   694: 'Spare_Fault_694', class No Acknowledgement, trigger "DB302_HMI_Faults_Carrier10_Faults_3" bit 5
   695: 'Spare_Fault_695', class No Acknowledgement, trigger "DB302_HMI_Faults_Carrier10_Faults_3" bit 6
   696: 'Spare_Fault_696', class No Acknowledgement, trigger "DB302_HMI_Faults_Carrier10_Faults_3" bit 7
   697: 'Spare_Fault_697', class No Acknowledgement, trigger "DB302_HMI_Faults_Carrier10_Faults_3" bit 8
   698: 'Spare_Fault_698', class No Acknowledgement, trigger "DB302_HMI_Faults_Carrier10_Faults_3" bit 9
   699: 'Spare_Fault_699', class No Acknowledgement, trigger "DB302_HMI_Faults_Carrier10_Faults_3" bit 10
   700: 'Spare_Fault_700', class No Acknowledgement, trigger "DB302_HMI_Faults_Carrier10_Faults_3" bit 11
   701: 'Spare_Fault_701', class No Acknowledgement, trigger "DB302_HMI_Faults_Carrier10_Faults_3" bit 12
   702: 'Spare_Fault_702', class No Acknowledgement, trigger "DB302_HMI_Faults_Carrier10_Faults_3" bit 13
   703: 'Spare_Fault_703', class No Acknowledgement, trigger "DB302_HMI_Faults_Carrier10_Faults_3" bit 14
   704: 'Spare_Fault_704', class No Acknowledgement, trigger "DB302_HMI_Faults_Carrier10_Faults_3" bit 15
   705: 'Carrier 11 Disconnect Open Power Fault DI11.0', class No Acknowledgement, trigger "DB302_HMI_Faults_Carrier11_Faults_0" bit 0
   706: 'Carrier 11 Drive Profinet Comm Fault', class No Acknowledgement, trigger "DB302_HMI_Faults_Carrier11_Faults_0" bit 1
   707: 'Carrier 11 Production Stop Not Reset', class No Acknowledgement, trigger "DB302_HMI_Faults_Carrier11_Faults_0" bit 2
   708: 'Carrier 11 CB02122 Tripped', class No Acknowledgement, trigger "DB302_HMI_Faults_Carrier11_Faults_0" bit 3
   709: 'Carrier 11 CB02123 Tripped', class No Acknowledgement, trigger "DB302_HMI_Faults_Carrier11_Faults_0" bit 4
   710: 'Carrier 11 AUX1 CB Tripped', class No Acknowledgement, trigger "DB302_HMI_Faults_Carrier11_Faults_0" bit 5
   711: 'Carrier 11 AUX2 CB Tripped', class No Acknowledgement, trigger "DB302_HMI_Faults_Carrier11_Faults_0" bit 6
   712: 'Carrier 11 PLC Not Communicating', class No Acknowledgement, trigger "DB302_HMI_Faults_Carrier11_Faults_0" bit 7
   713: 'Carrier 11 Safe Input Card Fault', class No Acknowledgement, trigger "DB302_HMI_Faults_Carrier11_Faults_0" bit 8
   714: 'Carrier 11 Safe Output Card Fault', class No Acknowledgement, trigger "DB302_HMI_Faults_Carrier11_Faults_0" bit 9
   715: 'Carrier 11 Standard Input Card Fault', class No Acknowledgement, trigger "DB302_HMI_Faults_Carrier11_Faults_0" bit 10
   716: 'Carrier 11 Standard Output Card Fault', class No Acknowledgement, trigger "DB302_HMI_Faults_Carrier11_Faults_0" bit 11
   717: 'Carrier 11 Encoder Position Fault', class No Acknowledgement, trigger "DB302_HMI_Faults_Carrier11_Faults_0" bit 12
   718: 'Carrier 11 Encoder Internal Error', class No Acknowledgement, trigger "DB302_HMI_Faults_Carrier11_Faults_0" bit 13
   719: 'Carrier 11 Encoder Comm Fault', class No Acknowledgement, trigger "DB302_HMI_Faults_Carrier11_Faults_0" bit 14
   720: 'Carrier 11 HMI Comm Fault', class No Acknowledgement, trigger "DB302_HMI_Faults_Carrier11_Faults_0" bit 15
   721: 'Carrier 11 Crash Detection Fault', class No Acknowledgement, trigger "DB302_HMI_Faults_Carrier11_Faults_1" bit 0
   722: 'Carrier 11 Carrier Number Invalid', class No Acknowledgement, trigger "DB302_HMI_Faults_Carrier11_Faults_1" bit 1
   723: 'Carrier 11 Drive: PROFINET configuration error', class No Acknowledgement, trigger "DB302_HMI_Faults_Carrier11_Faults_1" bit 2
   724: 'Carrier 11 Drive: Error internal communications', class No Acknowledgement, trigger "DB302_HMI_Faults_Carrier11_Faults_1" bit 3
   725: 'Carrier 11 Drive: Motor overtemperature', class No Acknowledgement, trigger "DB302_HMI_Faults_Carrier11_Faults_1" bit 4
   726: 'Carrier 11 Drive: Motor overcurrent', class No Acknowledgement, trigger "DB302_HMI_Faults_Carrier11_Faults_1" bit 5
   727: 'Carrier 11 Drive: Infeed or power unit not ready', class No Acknowledgement, trigger "DB302_HMI_Faults_Carrier11_Faults_1" bit 6
   728: 'Carrier 11 Drive: Short-circuit/ground fault detected', class No Acknowledgement, trigger "DB302_HMI_Faults_Carrier11_Faults_1" bit 7
   729: 'Carrier 11 Drive: PROFINET Setpoint timeout', class No Acknowledgement, trigger "DB302_HMI_Faults_Carrier11_Faults_1" bit 8
   730: 'Carrier 11 Power unit: Overcurrent', class No Acknowledgement, trigger "DB302_HMI_Faults_Carrier11_Faults_1" bit 9
   731: 'Carrier 11 Power unit: DC link voltage overvoltage', class No Acknowledgement, trigger "DB302_HMI_Faults_Carrier11_Faults_1" bit 10
   732: 'Carrier 11 Power unit: DC link voltage undervoltage', class No Acknowledgement, trigger "DB302_HMI_Faults_Carrier11_Faults_1" bit 11
   733: 'Carrier 11 Power unit: Line phase failure in main circuit', class No Acknowledgement, trigger "DB302_HMI_Faults_Carrier11_Faults_1" bit 12
   734: 'Carrier 11 Power unit: Phase failure motor cable', class No Acknowledgement, trigger "DB302_HMI_Faults_Carrier11_Faults_1" bit 13
   735: 'Carrier 11 Power unit: Ground fault', class No Acknowledgement, trigger "DB302_HMI_Faults_Carrier11_Faults_1" bit 14
   736: 'Spare_Fault_736', class No Acknowledgement, trigger "DB302_HMI_Faults_Carrier11_Faults_1" bit 15
   737: 'Carrier 11 Motion Off Fault', class No Acknowledgement, trigger "DB302_HMI_Faults_Carrier11_Faults_2" bit 0
   738: 'Carrier 11 Motion On Fault', class No Acknowledgement, trigger "DB302_HMI_Faults_Carrier11_Faults_2" bit 1
   739: 'Carrier 11 Spacing Fault', class No Acknowledgement, trigger "DB302_HMI_Faults_Carrier11_Faults_2" bit 2
   740: 'Carrier 11 Duplicate Carrier Number Fault', class No Acknowledgement, trigger "DB302_HMI_Faults_Carrier11_Faults_2" bit 3
   741: 'Spare_Fault_741', class No Acknowledgement, trigger "DB302_HMI_Faults_Carrier11_Faults_2" bit 4
   742: 'Spare_Fault_742', class No Acknowledgement, trigger "DB302_HMI_Faults_Carrier11_Faults_2" bit 5
   743: 'Spare_Fault_743', class No Acknowledgement, trigger "DB302_HMI_Faults_Carrier11_Faults_2" bit 6
   744: 'Spare_Fault_744', class No Acknowledgement, trigger "DB302_HMI_Faults_Carrier11_Faults_2" bit 7
   745: 'Spare_Fault_745', class No Acknowledgement, trigger "DB302_HMI_Faults_Carrier11_Faults_2" bit 8
   746: 'Spare_Fault_746', class No Acknowledgement, trigger "DB302_HMI_Faults_Carrier11_Faults_2" bit 9
   747: 'Spare_Fault_747', class No Acknowledgement, trigger "DB302_HMI_Faults_Carrier11_Faults_2" bit 10
   748: 'Spare_Fault_748', class No Acknowledgement, trigger "DB302_HMI_Faults_Carrier11_Faults_2" bit 11
   749: 'Spare_Fault_749', class No Acknowledgement, trigger "DB302_HMI_Faults_Carrier11_Faults_2" bit 12
   750: 'Spare_Fault_750', class No Acknowledgement, trigger "DB302_HMI_Faults_Carrier11_Faults_2" bit 13
   751: 'Spare_Fault_751', class No Acknowledgement, trigger "DB302_HMI_Faults_Carrier11_Faults_2" bit 14
   752: 'Spare_Fault_752', class No Acknowledgement, trigger "DB302_HMI_Faults_Carrier11_Faults_2" bit 15
   753: 'Spare_Fault_753', class No Acknowledgement, trigger "DB302_HMI_Faults_Carrier11_Faults_3" bit 0
   754: 'Spare_Fault_754', class No Acknowledgement, trigger "DB302_HMI_Faults_Carrier11_Faults_3" bit 1
   755: 'Spare_Fault_755', class No Acknowledgement, trigger "DB302_HMI_Faults_Carrier11_Faults_3" bit 2
   756: 'Spare_Fault_756', class No Acknowledgement, trigger "DB302_HMI_Faults_Carrier11_Faults_3" bit 3
   757: 'Spare_Fault_757', class No Acknowledgement, trigger "DB302_HMI_Faults_Carrier11_Faults_3" bit 4
   758: 'Spare_Fault_758', class No Acknowledgement, trigger "DB302_HMI_Faults_Carrier11_Faults_3" bit 5
   759: 'Spare_Fault_759', class No Acknowledgement, trigger "DB302_HMI_Faults_Carrier11_Faults_3" bit 6
   760: 'Spare_Fault_760', class No Acknowledgement, trigger "DB302_HMI_Faults_Carrier11_Faults_3" bit 7
   761: 'Spare_Fault_761', class No Acknowledgement, trigger "DB302_HMI_Faults_Carrier11_Faults_3" bit 8
   762: 'Spare_Fault_762', class No Acknowledgement, trigger "DB302_HMI_Faults_Carrier11_Faults_3" bit 9
   763: 'Spare_Fault_763', class No Acknowledgement, trigger "DB302_HMI_Faults_Carrier11_Faults_3" bit 10
   764: 'Spare_Fault_764', class No Acknowledgement, trigger "DB302_HMI_Faults_Carrier11_Faults_3" bit 11
   765: 'Spare_Fault_765', class No Acknowledgement, trigger "DB302_HMI_Faults_Carrier11_Faults_3" bit 12
   766: 'Spare_Fault_766', class No Acknowledgement, trigger "DB302_HMI_Faults_Carrier11_Faults_3" bit 13
   767: 'Spare_Fault_767', class No Acknowledgement, trigger "DB302_HMI_Faults_Carrier11_Faults_3" bit 14
   768: 'Spare_Fault_768', class No Acknowledgement, trigger "DB302_HMI_Faults_Carrier11_Faults_3" bit 15
   769: 'Carrier 12 Disconnect Open Power Fault DI11.0', class No Acknowledgement, trigger "DB302_HMI_Faults_Carrier12_Faults_0" bit 0
   770: 'Carrier 12 Drive Profinet Comm Fault', class No Acknowledgement, trigger "DB302_HMI_Faults_Carrier12_Faults_0" bit 1
   771: 'Carrier 12 Production Stop Not Reset', class No Acknowledgement, trigger "DB302_HMI_Faults_Carrier12_Faults_0" bit 2
   772: 'Carrier 12 CB02122 Tripped', class No Acknowledgement, trigger "DB302_HMI_Faults_Carrier12_Faults_0" bit 3
   773: 'Carrier 12 CB02123 Tripped', class No Acknowledgement, trigger "DB302_HMI_Faults_Carrier12_Faults_0" bit 4
   774: 'Carrier 12 AUX1 CB Tripped', class No Acknowledgement, trigger "DB302_HMI_Faults_Carrier12_Faults_0" bit 5
   775: 'Carrier 12 AUX2 CB Tripped', class No Acknowledgement, trigger "DB302_HMI_Faults_Carrier12_Faults_0" bit 6
   776: 'Carrier 12 PLC Not Communicating', class No Acknowledgement, trigger "DB302_HMI_Faults_Carrier12_Faults_0" bit 7
   777: 'Carrier 12 Safe Input Card Fault', class No Acknowledgement, trigger "DB302_HMI_Faults_Carrier12_Faults_0" bit 8
   778: 'Carrier 12 Safe Output Card Fault', class No Acknowledgement, trigger "DB302_HMI_Faults_Carrier12_Faults_0" bit 9
   779: 'Carrier 12 Standard Input Card Fault', class No Acknowledgement, trigger "DB302_HMI_Faults_Carrier12_Faults_0" bit 10
   780: 'Carrier 12 Standard Output Card Fault', class No Acknowledgement, trigger "DB302_HMI_Faults_Carrier12_Faults_0" bit 11
   781: 'Carrier 12 Encoder Position Fault', class No Acknowledgement, trigger "DB302_HMI_Faults_Carrier12_Faults_0" bit 12
   782: 'Carrier 12 Encoder Internal Error', class No Acknowledgement, trigger "DB302_HMI_Faults_Carrier12_Faults_0" bit 13
   783: 'Carrier 12 Encoder Comm Fault', class No Acknowledgement, trigger "DB302_HMI_Faults_Carrier12_Faults_0" bit 14
   784: 'Carrier 12 HMI Comm Fault', class No Acknowledgement, trigger "DB302_HMI_Faults_Carrier12_Faults_0" bit 15
   785: 'Carrier 12 Crash Detection Fault', class No Acknowledgement, trigger "DB302_HMI_Faults_Carrier12_Faults_1" bit 0
   786: 'Carrier 12 Carrier Number Invalid', class No Acknowledgement, trigger "DB302_HMI_Faults_Carrier12_Faults_1" bit 1
   787: 'Carrier 12 Drive: PROFINET configuration error', class No Acknowledgement, trigger "DB302_HMI_Faults_Carrier12_Faults_1" bit 2
   788: 'Carrier 12 Drive: Error internal communications', class No Acknowledgement, trigger "DB302_HMI_Faults_Carrier12_Faults_1" bit 3
   789: 'Carrier 12 Drive: Motor overtemperature', class No Acknowledgement, trigger "DB302_HMI_Faults_Carrier12_Faults_1" bit 4
   790: 'Carrier 12 Drive: Motor overcurrent', class No Acknowledgement, trigger "DB302_HMI_Faults_Carrier12_Faults_1" bit 5
   791: 'Carrier 12 Drive: Infeed or power unit not ready', class No Acknowledgement, trigger "DB302_HMI_Faults_Carrier12_Faults_1" bit 6
   792: 'Carrier 12 Drive: Short-circuit/ground fault detected', class No Acknowledgement, trigger "DB302_HMI_Faults_Carrier12_Faults_1" bit 7
   793: 'Carrier 12 Drive: PROFINET Setpoint timeout', class No Acknowledgement, trigger "DB302_HMI_Faults_Carrier12_Faults_1" bit 8
   794: 'Carrier 12 Power unit: Overcurrent', class No Acknowledgement, trigger "DB302_HMI_Faults_Carrier12_Faults_1" bit 9
   795: 'Carrier 12 Power unit: DC link voltage overvoltage', class No Acknowledgement, trigger "DB302_HMI_Faults_Carrier12_Faults_1" bit 10
   796: 'Carrier 12 Power unit: DC link voltage undervoltage', class No Acknowledgement, trigger "DB302_HMI_Faults_Carrier12_Faults_1" bit 11
   797: 'Carrier 12 Power unit: Line phase failure in main circuit', class No Acknowledgement, trigger "DB302_HMI_Faults_Carrier12_Faults_1" bit 12
   798: 'Carrier 12 Power unit: Phase failure motor cable', class No Acknowledgement, trigger "DB302_HMI_Faults_Carrier12_Faults_1" bit 13
   799: 'Carrier 12 Power unit: Ground fault', class No Acknowledgement, trigger "DB302_HMI_Faults_Carrier12_Faults_1" bit 14
   800: 'Spare_Fault_800', class No Acknowledgement, trigger "DB302_HMI_Faults_Carrier12_Faults_1" bit 15
   801: 'Carrier 12 Motion Off Fault', class No Acknowledgement, trigger "DB302_HMI_Faults_Carrier12_Faults_2" bit 0
   802: 'Carrier 12 Motion On Fault', class No Acknowledgement, trigger "DB302_HMI_Faults_Carrier12_Faults_2" bit 1
   803: 'Carrier 12 Spacing Fault', class No Acknowledgement, trigger "DB302_HMI_Faults_Carrier12_Faults_2" bit 2
   804: 'Carrier 12 Duplicate Carrier Number Fault', class No Acknowledgement, trigger "DB302_HMI_Faults_Carrier12_Faults_2" bit 3
   805: 'Spare_Fault_805', class No Acknowledgement, trigger "DB302_HMI_Faults_Carrier12_Faults_2" bit 4
   806: 'Spare_Fault_806', class No Acknowledgement, trigger "DB302_HMI_Faults_Carrier12_Faults_2" bit 5
   807: 'Spare_Fault_807', class No Acknowledgement, trigger "DB302_HMI_Faults_Carrier12_Faults_2" bit 6
   808: 'Spare_Fault_808', class No Acknowledgement, trigger "DB302_HMI_Faults_Carrier12_Faults_2" bit 7
   809: 'Spare_Fault_809', class No Acknowledgement, trigger "DB302_HMI_Faults_Carrier12_Faults_2" bit 8
   810: 'Spare_Fault_810', class No Acknowledgement, trigger "DB302_HMI_Faults_Carrier12_Faults_2" bit 9
   811: 'Spare_Fault_811', class No Acknowledgement, trigger "DB302_HMI_Faults_Carrier12_Faults_2" bit 10
   812: 'Spare_Fault_812', class No Acknowledgement, trigger "DB302_HMI_Faults_Carrier12_Faults_2" bit 11
   813: 'Spare_Fault_813', class No Acknowledgement, trigger "DB302_HMI_Faults_Carrier12_Faults_2" bit 12
   814: 'Spare_Fault_814', class No Acknowledgement, trigger "DB302_HMI_Faults_Carrier12_Faults_2" bit 13
   815: 'Spare_Fault_815', class No Acknowledgement, trigger "DB302_HMI_Faults_Carrier12_Faults_2" bit 14
   816: 'Spare_Fault_816', class No Acknowledgement, trigger "DB302_HMI_Faults_Carrier12_Faults_2" bit 15
   817: 'Spare_Fault_817', class No Acknowledgement, trigger "DB302_HMI_Faults_Carrier12_Faults_3" bit 0
   818: 'Spare_Fault_818', class No Acknowledgement, trigger "DB302_HMI_Faults_Carrier12_Faults_3" bit 1
   819: 'Spare_Fault_819', class No Acknowledgement, trigger "DB302_HMI_Faults_Carrier12_Faults_3" bit 2
   820: 'Spare_Fault_820', class No Acknowledgement, trigger "DB302_HMI_Faults_Carrier12_Faults_3" bit 3
   821: 'Spare_Fault_821', class No Acknowledgement, trigger "DB302_HMI_Faults_Carrier12_Faults_3" bit 4
   822: 'Spare_Fault_822', class No Acknowledgement, trigger "DB302_HMI_Faults_Carrier12_Faults_3" bit 5
   823: 'Spare_Fault_823', class No Acknowledgement, trigger "DB302_HMI_Faults_Carrier12_Faults_3" bit 6
   824: 'Spare_Fault_824', class No Acknowledgement, trigger "DB302_HMI_Faults_Carrier12_Faults_3" bit 7
   825: 'Spare_Fault_825', class No Acknowledgement, trigger "DB302_HMI_Faults_Carrier12_Faults_3" bit 8
   826: 'Spare_Fault_826', class No Acknowledgement, trigger "DB302_HMI_Faults_Carrier12_Faults_3" bit 9
   827: 'Spare_Fault_827', class No Acknowledgement, trigger "DB302_HMI_Faults_Carrier12_Faults_3" bit 10
   828: 'Spare_Fault_828', class No Acknowledgement, trigger "DB302_HMI_Faults_Carrier12_Faults_3" bit 11
   829: 'Spare_Fault_829', class No Acknowledgement, trigger "DB302_HMI_Faults_Carrier12_Faults_3" bit 12
   830: 'Spare_Fault_830', class No Acknowledgement, trigger "DB302_HMI_Faults_Carrier12_Faults_3" bit 13
   831: 'Spare_Fault_831', class No Acknowledgement, trigger "DB302_HMI_Faults_Carrier12_Faults_3" bit 14
   832: 'Spare_Fault_832', class No Acknowledgement, trigger "DB302_HMI_Faults_Carrier12_Faults_3" bit 15
   833: 'Carrier 13 Disconnect Open Power Fault DI11.0', class No Acknowledgement, trigger "DB302_HMI_Faults_Carrier13_Faults_0" bit 0
   834: 'Carrier 13 Drive Profinet Comm Fault', class No Acknowledgement, trigger "DB302_HMI_Faults_Carrier13_Faults_0" bit 1
   835: 'Carrier 13 Production Stop Not Reset', class No Acknowledgement, trigger "DB302_HMI_Faults_Carrier13_Faults_0" bit 2
   836: 'Carrier 13 CB02122 Tripped', class No Acknowledgement, trigger "DB302_HMI_Faults_Carrier13_Faults_0" bit 3
   837: 'Carrier 13 CB02123 Tripped', class No Acknowledgement, trigger "DB302_HMI_Faults_Carrier13_Faults_0" bit 4
   838: 'Carrier 13 AUX1 CB Tripped', class No Acknowledgement, trigger "DB302_HMI_Faults_Carrier13_Faults_0" bit 5
   839: 'Carrier 13 AUX2 CB Tripped', class No Acknowledgement, trigger "DB302_HMI_Faults_Carrier13_Faults_0" bit 6
   840: 'Carrier 13 PLC Not Communicating', class No Acknowledgement, trigger "DB302_HMI_Faults_Carrier13_Faults_0" bit 7
   841: 'Carrier 13 Safe Input Card Fault', class No Acknowledgement, trigger "DB302_HMI_Faults_Carrier13_Faults_0" bit 8
   842: 'Carrier 13 Safe Output Card Fault', class No Acknowledgement, trigger "DB302_HMI_Faults_Carrier13_Faults_0" bit 9
   843: 'Carrier 13 Standard Input Card Fault', class No Acknowledgement, trigger "DB302_HMI_Faults_Carrier13_Faults_0" bit 10
   844: 'Carrier 13 Standard Output Card Fault', class No Acknowledgement, trigger "DB302_HMI_Faults_Carrier13_Faults_0" bit 11
   845: 'Carrier 13 Encoder Position Fault', class No Acknowledgement, trigger "DB302_HMI_Faults_Carrier13_Faults_0" bit 12
   846: 'Carrier 13 Encoder Internal Error', class No Acknowledgement, trigger "DB302_HMI_Faults_Carrier13_Faults_0" bit 13
   847: 'Carrier 13 Encoder Comm Fault', class No Acknowledgement, trigger "DB302_HMI_Faults_Carrier13_Faults_0" bit 14
   848: 'Carrier 13 HMI Comm Fault', class No Acknowledgement, trigger "DB302_HMI_Faults_Carrier13_Faults_0" bit 15
   849: 'Carrier 13 Crash Detection Fault', class No Acknowledgement, trigger "DB302_HMI_Faults_Carrier13_Faults_1" bit 0
   850: 'Carrier 13 Carrier Number Invalid', class No Acknowledgement, trigger "DB302_HMI_Faults_Carrier13_Faults_1" bit 1
   851: 'Carrier 13 Drive: PROFINET configuration error', class No Acknowledgement, trigger "DB302_HMI_Faults_Carrier13_Faults_1" bit 2
   852: 'Carrier 13 Drive: Error internal communications', class No Acknowledgement, trigger "DB302_HMI_Faults_Carrier13_Faults_1" bit 3
   853: 'Carrier 13 Drive: Motor overtemperature', class No Acknowledgement, trigger "DB302_HMI_Faults_Carrier13_Faults_1" bit 4
   854: 'Carrier 13 Drive: Motor overcurrent', class No Acknowledgement, trigger "DB302_HMI_Faults_Carrier13_Faults_1" bit 5
   855: 'Carrier 13 Drive: Infeed or power unit not ready', class No Acknowledgement, trigger "DB302_HMI_Faults_Carrier13_Faults_1" bit 6
   856: 'Carrier 13 Drive: Short-circuit/ground fault detected', class No Acknowledgement, trigger "DB302_HMI_Faults_Carrier13_Faults_1" bit 7
   857: 'Carrier 13 Drive: PROFINET Setpoint timeout', class No Acknowledgement, trigger "DB302_HMI_Faults_Carrier13_Faults_1" bit 8
   858: 'Carrier 13 Power unit: Overcurrent', class No Acknowledgement, trigger "DB302_HMI_Faults_Carrier13_Faults_1" bit 9
   859: 'Carrier 13 Power unit: DC link voltage overvoltage', class No Acknowledgement, trigger "DB302_HMI_Faults_Carrier13_Faults_1" bit 10
   860: 'Carrier 13 Power unit: DC link voltage undervoltage', class No Acknowledgement, trigger "DB302_HMI_Faults_Carrier13_Faults_1" bit 11
   861: 'Carrier 13 Power unit: Line phase failure in main circuit', class No Acknowledgement, trigger "DB302_HMI_Faults_Carrier13_Faults_1" bit 12
   862: 'Carrier 13 Power unit: Phase failure motor cable', class No Acknowledgement, trigger "DB302_HMI_Faults_Carrier13_Faults_1" bit 13
   863: 'Carrier 13 Power unit: Ground fault', class No Acknowledgement, trigger "DB302_HMI_Faults_Carrier13_Faults_1" bit 14
   864: 'Spare_Fault_864', class No Acknowledgement, trigger "DB302_HMI_Faults_Carrier13_Faults_1" bit 15
   865: 'Carrier 13 Motion Off Fault', class No Acknowledgement, trigger "DB302_HMI_Faults_Carrier13_Faults_2" bit 0
   866: 'Carrier 13 Motion On Fault', class No Acknowledgement, trigger "DB302_HMI_Faults_Carrier13_Faults_2" bit 1
   867: 'Carrier 13 Spacing Fault', class No Acknowledgement, trigger "DB302_HMI_Faults_Carrier13_Faults_2" bit 2
   868: 'Carrier 13 Duplicate Carrier Number Fault', class No Acknowledgement, trigger "DB302_HMI_Faults_Carrier13_Faults_2" bit 3
   869: 'Spare_Fault_869', class No Acknowledgement, trigger "DB302_HMI_Faults_Carrier13_Faults_2" bit 4
   870: 'Spare_Fault_870', class No Acknowledgement, trigger "DB302_HMI_Faults_Carrier13_Faults_2" bit 5
   871: 'Spare_Fault_871', class No Acknowledgement, trigger "DB302_HMI_Faults_Carrier13_Faults_2" bit 6
   872: 'Spare_Fault_872', class No Acknowledgement, trigger "DB302_HMI_Faults_Carrier13_Faults_2" bit 7
   873: 'Spare_Fault_873', class No Acknowledgement, trigger "DB302_HMI_Faults_Carrier13_Faults_2" bit 8
   874: 'Spare_Fault_874', class No Acknowledgement, trigger "DB302_HMI_Faults_Carrier13_Faults_2" bit 9
   875: 'Spare_Fault_875', class No Acknowledgement, trigger "DB302_HMI_Faults_Carrier13_Faults_2" bit 10
   876: 'Spare_Fault_876', class No Acknowledgement, trigger "DB302_HMI_Faults_Carrier13_Faults_2" bit 11
   877: 'Spare_Fault_877', class No Acknowledgement, trigger "DB302_HMI_Faults_Carrier13_Faults_2" bit 12
   878: 'Spare_Fault_878', class No Acknowledgement, trigger "DB302_HMI_Faults_Carrier13_Faults_2" bit 13
   879: 'Spare_Fault_879', class No Acknowledgement, trigger "DB302_HMI_Faults_Carrier13_Faults_2" bit 14
   880: 'Spare_Fault_880', class No Acknowledgement, trigger "DB302_HMI_Faults_Carrier13_Faults_2" bit 15
   881: 'Spare_Fault_881', class No Acknowledgement, trigger "DB302_HMI_Faults_Carrier13_Faults_3" bit 0
   882: 'Spare_Fault_882', class No Acknowledgement, trigger "DB302_HMI_Faults_Carrier13_Faults_3" bit 1
   883: 'Spare_Fault_883', class No Acknowledgement, trigger "DB302_HMI_Faults_Carrier13_Faults_3" bit 2
   884: 'Spare_Fault_884', class No Acknowledgement, trigger "DB302_HMI_Faults_Carrier13_Faults_3" bit 3
   885: 'Spare_Fault_885', class No Acknowledgement, trigger "DB302_HMI_Faults_Carrier13_Faults_3" bit 4
   886: 'Spare_Fault_886', class No Acknowledgement, trigger "DB302_HMI_Faults_Carrier13_Faults_3" bit 5
   887: 'Spare_Fault_887', class No Acknowledgement, trigger "DB302_HMI_Faults_Carrier13_Faults_3" bit 6
   888: 'Spare_Fault_888', class No Acknowledgement, trigger "DB302_HMI_Faults_Carrier13_Faults_3" bit 7
   889: 'Spare_Fault_889', class No Acknowledgement, trigger "DB302_HMI_Faults_Carrier13_Faults_3" bit 8
   890: 'Spare_Fault_890', class No Acknowledgement, trigger "DB302_HMI_Faults_Carrier13_Faults_3" bit 9
   891: 'Spare_Fault_891', class No Acknowledgement, trigger "DB302_HMI_Faults_Carrier13_Faults_3" bit 10
   892: 'Spare_Fault_892', class No Acknowledgement, trigger "DB302_HMI_Faults_Carrier13_Faults_3" bit 11
   893: 'Spare_Fault_893', class No Acknowledgement, trigger "DB302_HMI_Faults_Carrier13_Faults_3" bit 12
   894: 'Spare_Fault_894', class No Acknowledgement, trigger "DB302_HMI_Faults_Carrier13_Faults_3" bit 13
   895: 'Spare_Fault_895', class No Acknowledgement, trigger "DB302_HMI_Faults_Carrier13_Faults_3" bit 14
   896: 'Spare_Fault_896', class No Acknowledgement, trigger "DB302_HMI_Faults_Carrier13_Faults_3" bit 15
   897: 'Carrier 14 Disconnect Open Power Fault DI11.0', class No Acknowledgement, trigger "DB302_HMI_Faults_Carrier14_Faults_0" bit 0
   898: 'Carrier 14 Drive Profinet Comm Fault', class No Acknowledgement, trigger "DB302_HMI_Faults_Carrier14_Faults_0" bit 1
   899: 'Carrier 14 Production Stop Not Reset', class No Acknowledgement, trigger "DB302_HMI_Faults_Carrier14_Faults_0" bit 2
   900: 'Carrier 14 CB02122 Tripped', class No Acknowledgement, trigger "DB302_HMI_Faults_Carrier14_Faults_0" bit 3
   901: 'Carrier 14 CB02123 Tripped', class No Acknowledgement, trigger "DB302_HMI_Faults_Carrier14_Faults_0" bit 4
   902: 'Carrier 14 AUX1 CB Tripped', class No Acknowledgement, trigger "DB302_HMI_Faults_Carrier14_Faults_0" bit 5
   903: 'Carrier 14 AUX2 CB Tripped', class No Acknowledgement, trigger "DB302_HMI_Faults_Carrier14_Faults_0" bit 6
   904: 'Carrier 14 PLC Not Communicating', class No Acknowledgement, trigger "DB302_HMI_Faults_Carrier14_Faults_0" bit 7
   905: 'Carrier 14 Safe Input Card Fault', class No Acknowledgement, trigger "DB302_HMI_Faults_Carrier14_Faults_0" bit 8
   906: 'Carrier 14 Safe Output Card Fault', class No Acknowledgement, trigger "DB302_HMI_Faults_Carrier14_Faults_0" bit 9
   907: 'Carrier 14 Standard Input Card Fault', class No Acknowledgement, trigger "DB302_HMI_Faults_Carrier14_Faults_0" bit 10
   908: 'Carrier 14 Standard Output Card Fault', class No Acknowledgement, trigger "DB302_HMI_Faults_Carrier14_Faults_0" bit 11
   909: 'Carrier 14 Encoder Position Fault', class No Acknowledgement, trigger "DB302_HMI_Faults_Carrier14_Faults_0" bit 12
   910: 'Carrier 14 Encoder Internal Error', class No Acknowledgement, trigger "DB302_HMI_Faults_Carrier14_Faults_0" bit 13
   911: 'Carrier 14 Encoder Comm Fault', class No Acknowledgement, trigger "DB302_HMI_Faults_Carrier14_Faults_0" bit 14
   912: 'Carrier 14 HMI Comm Fault', class No Acknowledgement, trigger "DB302_HMI_Faults_Carrier14_Faults_0" bit 15
   913: 'Carrier 14 Crash Detection Fault', class No Acknowledgement, trigger "DB302_HMI_Faults_Carrier14_Faults_1" bit 0
   914: 'Carrier 14 Carrier Number Invalid', class No Acknowledgement, trigger "DB302_HMI_Faults_Carrier14_Faults_1" bit 1
   915: 'Carrier 14 Drive: PROFINET configuration error', class No Acknowledgement, trigger "DB302_HMI_Faults_Carrier14_Faults_1" bit 2
   916: 'Carrier 14 Drive: Error internal communications', class No Acknowledgement, trigger "DB302_HMI_Faults_Carrier14_Faults_1" bit 3
   917: 'Carrier 14 Drive: Motor overtemperature', class No Acknowledgement, trigger "DB302_HMI_Faults_Carrier14_Faults_1" bit 4
   918: 'Carrier 14 Drive: Motor overcurrent', class No Acknowledgement, trigger "DB302_HMI_Faults_Carrier14_Faults_1" bit 5
   919: 'Carrier 14 Drive: Infeed or power unit not ready', class No Acknowledgement, trigger "DB302_HMI_Faults_Carrier14_Faults_1" bit 6
   920: 'Carrier 14 Drive: Short-circuit/ground fault detected', class No Acknowledgement, trigger "DB302_HMI_Faults_Carrier14_Faults_1" bit 7
   921: 'Carrier 14 Drive: PROFINET Setpoint timeout', class No Acknowledgement, trigger "DB302_HMI_Faults_Carrier14_Faults_1" bit 8
   922: 'Carrier 14 Power unit: Overcurrent', class No Acknowledgement, trigger "DB302_HMI_Faults_Carrier14_Faults_1" bit 9
   923: 'Carrier 14 Power unit: DC link voltage overvoltage', class No Acknowledgement, trigger "DB302_HMI_Faults_Carrier14_Faults_1" bit 10
   924: 'Carrier 14 Power unit: DC link voltage undervoltage', class No Acknowledgement, trigger "DB302_HMI_Faults_Carrier14_Faults_1" bit 11
   925: 'Carrier 14 Power unit: Line phase failure in main circuit', class No Acknowledgement, trigger "DB302_HMI_Faults_Carrier14_Faults_1" bit 12
   926: 'Carrier 14 Power unit: Phase failure motor cable', class No Acknowledgement, trigger "DB302_HMI_Faults_Carrier14_Faults_1" bit 13
   927: 'Carrier 14 Power unit: Ground fault', class No Acknowledgement, trigger "DB302_HMI_Faults_Carrier14_Faults_1" bit 14
   928: 'Spare_Fault_928', class No Acknowledgement, trigger "DB302_HMI_Faults_Carrier14_Faults_1" bit 15
   929: 'Carrier 14 Motion Off Fault', class No Acknowledgement, trigger "DB302_HMI_Faults_Carrier14_Faults_2" bit 0
   930: 'Carrier 14 Motion On Fault', class No Acknowledgement, trigger "DB302_HMI_Faults_Carrier14_Faults_2" bit 1
   931: 'Carrier 14 Spacing Fault', class No Acknowledgement, trigger "DB302_HMI_Faults_Carrier14_Faults_2" bit 2
   932: 'Carrier 14 Duplicate Carrier Number Fault', class No Acknowledgement, trigger "DB302_HMI_Faults_Carrier14_Faults_2" bit 3
   933: 'Spare_Fault_933', class No Acknowledgement, trigger "DB302_HMI_Faults_Carrier14_Faults_2" bit 4
   934: 'Spare_Fault_934', class No Acknowledgement, trigger "DB302_HMI_Faults_Carrier14_Faults_2" bit 5
   935: 'Spare_Fault_935', class No Acknowledgement, trigger "DB302_HMI_Faults_Carrier14_Faults_2" bit 6
   936: 'Spare_Fault_936', class No Acknowledgement, trigger "DB302_HMI_Faults_Carrier14_Faults_2" bit 7
   937: 'Spare_Fault_937', class No Acknowledgement, trigger "DB302_HMI_Faults_Carrier14_Faults_2" bit 8
   938: 'Spare_Fault_938', class No Acknowledgement, trigger "DB302_HMI_Faults_Carrier14_Faults_2" bit 9
   939: 'Spare_Fault_939', class No Acknowledgement, trigger "DB302_HMI_Faults_Carrier14_Faults_2" bit 10
   940: 'Spare_Fault_940', class No Acknowledgement, trigger "DB302_HMI_Faults_Carrier14_Faults_2" bit 11
   941: 'Spare_Fault_941', class No Acknowledgement, trigger "DB302_HMI_Faults_Carrier14_Faults_2" bit 12
   942: 'Spare_Fault_942', class No Acknowledgement, trigger "DB302_HMI_Faults_Carrier14_Faults_2" bit 13
   943: 'Spare_Fault_943', class No Acknowledgement, trigger "DB302_HMI_Faults_Carrier14_Faults_2" bit 14
   944: 'Spare_Fault_944', class No Acknowledgement, trigger "DB302_HMI_Faults_Carrier14_Faults_2" bit 15
   945: 'Spare_Fault_945', class No Acknowledgement, trigger "DB302_HMI_Faults_Carrier14_Faults_3" bit 0
   946: 'Spare_Fault_946', class No Acknowledgement, trigger "DB302_HMI_Faults_Carrier14_Faults_3" bit 1
   947: 'Spare_Fault_947', class No Acknowledgement, trigger "DB302_HMI_Faults_Carrier14_Faults_3" bit 2
   948: 'Spare_Fault_948', class No Acknowledgement, trigger "DB302_HMI_Faults_Carrier14_Faults_3" bit 3
   949: 'Spare_Fault_949', class No Acknowledgement, trigger "DB302_HMI_Faults_Carrier14_Faults_3" bit 4
   950: 'Spare_Fault_950', class No Acknowledgement, trigger "DB302_HMI_Faults_Carrier14_Faults_3" bit 5
   951: 'Spare_Fault_951', class No Acknowledgement, trigger "DB302_HMI_Faults_Carrier14_Faults_3" bit 6
   952: 'Spare_Fault_952', class No Acknowledgement, trigger "DB302_HMI_Faults_Carrier14_Faults_3" bit 7
   953: 'Spare_Fault_953', class No Acknowledgement, trigger "DB302_HMI_Faults_Carrier14_Faults_3" bit 8
   954: 'Spare_Fault_954', class No Acknowledgement, trigger "DB302_HMI_Faults_Carrier14_Faults_3" bit 9
   955: 'Spare_Fault_955', class No Acknowledgement, trigger "DB302_HMI_Faults_Carrier14_Faults_3" bit 10
   956: 'Spare_Fault_956', class No Acknowledgement, trigger "DB302_HMI_Faults_Carrier14_Faults_3" bit 11
   957: 'Spare_Fault_957', class No Acknowledgement, trigger "DB302_HMI_Faults_Carrier14_Faults_3" bit 12
   958: 'Spare_Fault_958', class No Acknowledgement, trigger "DB302_HMI_Faults_Carrier14_Faults_3" bit 13
   959: 'Spare_Fault_959', class No Acknowledgement, trigger "DB302_HMI_Faults_Carrier14_Faults_3" bit 14
   960: 'Spare_Fault_960', class No Acknowledgement, trigger "DB302_HMI_Faults_Carrier14_Faults_3" bit 15
   961: 'Carrier 15 Disconnect Open Power Fault DI11.0', class No Acknowledgement, trigger "DB302_HMI_Faults_Carrier15_Faults_0" bit 0
   962: 'Carrier 15 Drive Profinet Comm Fault', class No Acknowledgement, trigger "DB302_HMI_Faults_Carrier15_Faults_0" bit 1
   963: 'Carrier 15 Production Stop Not Reset', class No Acknowledgement, trigger "DB302_HMI_Faults_Carrier15_Faults_0" bit 2
   964: 'Carrier 15 CB02122 Tripped', class No Acknowledgement, trigger "DB302_HMI_Faults_Carrier15_Faults_0" bit 3
   965: 'Carrier 15 CB02123 Tripped', class No Acknowledgement, trigger "DB302_HMI_Faults_Carrier15_Faults_0" bit 4
   966: 'Carrier 15 AUX1 CB Tripped', class No Acknowledgement, trigger "DB302_HMI_Faults_Carrier15_Faults_0" bit 5
   967: 'Carrier 15 AUX2 CB Tripped', class No Acknowledgement, trigger "DB302_HMI_Faults_Carrier15_Faults_0" bit 6
   968: 'Carrier 15 PLC Not Communicating', class No Acknowledgement, trigger "DB302_HMI_Faults_Carrier15_Faults_0" bit 7
   969: 'Carrier 15 Safe Input Card Fault', class No Acknowledgement, trigger "DB302_HMI_Faults_Carrier15_Faults_0" bit 8
   970: 'Carrier 15 Safe Output Card Fault', class No Acknowledgement, trigger "DB302_HMI_Faults_Carrier15_Faults_0" bit 9
   971: 'Carrier 15 Standard Input Card Fault', class No Acknowledgement, trigger "DB302_HMI_Faults_Carrier15_Faults_0" bit 10
   972: 'Carrier 15 Standard Output Card Fault', class No Acknowledgement, trigger "DB302_HMI_Faults_Carrier15_Faults_0" bit 11
   973: 'Carrier 15 Encoder Position Fault', class No Acknowledgement, trigger "DB302_HMI_Faults_Carrier15_Faults_0" bit 12
   974: 'Carrier 15 Encoder Internal Error', class No Acknowledgement, trigger "DB302_HMI_Faults_Carrier15_Faults_0" bit 13
   975: 'Carrier 15 Encoder Comm Fault', class No Acknowledgement, trigger "DB302_HMI_Faults_Carrier15_Faults_0" bit 14
   976: 'Carrier 15 HMI Comm Fault', class No Acknowledgement, trigger "DB302_HMI_Faults_Carrier15_Faults_0" bit 15
   977: 'Carrier 15 Crash Detection Fault', class No Acknowledgement, trigger "DB302_HMI_Faults_Carrier15_Faults_1" bit 0
   978: 'Carrier 15 Carrier Number Invalid', class No Acknowledgement, trigger "DB302_HMI_Faults_Carrier15_Faults_1" bit 1
   979: 'Carrier 15 Drive: PROFINET configuration error', class No Acknowledgement, trigger "DB302_HMI_Faults_Carrier15_Faults_1" bit 2
   980: 'Carrier 15 Drive: Error internal communications', class No Acknowledgement, trigger "DB302_HMI_Faults_Carrier15_Faults_1" bit 3
   981: 'Carrier 15 Drive: Motor overtemperature', class No Acknowledgement, trigger "DB302_HMI_Faults_Carrier15_Faults_1" bit 4
   982: 'Carrier 15 Drive: Motor overcurrent', class No Acknowledgement, trigger "DB302_HMI_Faults_Carrier15_Faults_1" bit 5
   983: 'Carrier 15 Drive: Infeed or power unit not ready', class No Acknowledgement, trigger "DB302_HMI_Faults_Carrier15_Faults_1" bit 6
   984: 'Carrier 15 Drive: Short-circuit/ground fault detected', class No Acknowledgement, trigger "DB302_HMI_Faults_Carrier15_Faults_1" bit 7
   985: 'Carrier 15 Drive: PROFINET Setpoint timeout', class No Acknowledgement, trigger "DB302_HMI_Faults_Carrier15_Faults_1" bit 8
   986: 'Carrier 15 Power unit: Overcurrent', class No Acknowledgement, trigger "DB302_HMI_Faults_Carrier15_Faults_1" bit 9
   987: 'Carrier 15 Power unit: DC link voltage overvoltage', class No Acknowledgement, trigger "DB302_HMI_Faults_Carrier15_Faults_1" bit 10
   988: 'Carrier 15 Power unit: DC link voltage undervoltage', class No Acknowledgement, trigger "DB302_HMI_Faults_Carrier15_Faults_1" bit 11
   989: 'Carrier 15 Power unit: Line phase failure in main circuit', class No Acknowledgement, trigger "DB302_HMI_Faults_Carrier15_Faults_1" bit 12
   990: 'Carrier 15 Power unit: Phase failure motor cable', class No Acknowledgement, trigger "DB302_HMI_Faults_Carrier15_Faults_1" bit 13
   991: 'Carrier 15 Power unit: Ground fault', class No Acknowledgement, trigger "DB302_HMI_Faults_Carrier15_Faults_1" bit 14
   992: 'Spare_Fault_992', class No Acknowledgement, trigger "DB302_HMI_Faults_Carrier15_Faults_1" bit 15
   993: 'Carrier 15 Motion Off Fault', class No Acknowledgement, trigger "DB302_HMI_Faults_Carrier15_Faults_2" bit 0
   994: 'Carrier 15 Motion On Fault', class No Acknowledgement, trigger "DB302_HMI_Faults_Carrier15_Faults_2" bit 1
   995: 'Carrier 15 Spacing Fault', class No Acknowledgement, trigger "DB302_HMI_Faults_Carrier15_Faults_2" bit 2
   996: 'Carrier 15 Duplicate Carrier Number Fault', class No Acknowledgement, trigger "DB302_HMI_Faults_Carrier15_Faults_2" bit 3
   997: 'Spare_Fault_997', class No Acknowledgement, trigger "DB302_HMI_Faults_Carrier15_Faults_2" bit 4
   998: 'Spare_Fault_998', class No Acknowledgement, trigger "DB302_HMI_Faults_Carrier15_Faults_2" bit 5
   999: 'Spare_Fault_999', class No Acknowledgement, trigger "DB302_HMI_Faults_Carrier15_Faults_2" bit 6
   1000: 'Spare_Fault_1000', class No Acknowledgement, trigger "DB302_HMI_Faults_Carrier15_Faults_2" bit 7
   1001: 'Spare_Fault_1001', class No Acknowledgement, trigger "DB302_HMI_Faults_Carrier15_Faults_2" bit 8
   1002: 'Spare_Fault_1002', class No Acknowledgement, trigger "DB302_HMI_Faults_Carrier15_Faults_2" bit 9
   1003: 'Spare_Fault_1003', class No Acknowledgement, trigger "DB302_HMI_Faults_Carrier15_Faults_2" bit 10
   1004: 'Spare_Fault_1004', class No Acknowledgement, trigger "DB302_HMI_Faults_Carrier15_Faults_2" bit 11
   1005: 'Spare_Fault_1005', class No Acknowledgement, trigger "DB302_HMI_Faults_Carrier15_Faults_2" bit 12
   1006: 'Spare_Fault_1006', class No Acknowledgement, trigger "DB302_HMI_Faults_Carrier15_Faults_2" bit 13
   1007: 'Spare_Fault_1007', class No Acknowledgement, trigger "DB302_HMI_Faults_Carrier15_Faults_2" bit 14
   1008: 'Spare_Fault_1008', class No Acknowledgement, trigger "DB302_HMI_Faults_Carrier15_Faults_2" bit 15
   1009: 'Spare_Fault_1009', class No Acknowledgement, trigger "DB302_HMI_Faults_Carrier15_Faults_3" bit 0
   1010: 'Spare_Fault_1010', class No Acknowledgement, trigger "DB302_HMI_Faults_Carrier15_Faults_3" bit 1
   1011: 'Spare_Fault_1011', class No Acknowledgement, trigger "DB302_HMI_Faults_Carrier15_Faults_3" bit 2
   1012: 'Spare_Fault_1012', class No Acknowledgement, trigger "DB302_HMI_Faults_Carrier15_Faults_3" bit 3
   1013: 'Spare_Fault_1013', class No Acknowledgement, trigger "DB302_HMI_Faults_Carrier15_Faults_3" bit 4
   1014: 'Spare_Fault_1014', class No Acknowledgement, trigger "DB302_HMI_Faults_Carrier15_Faults_3" bit 5
   1015: 'Spare_Fault_1015', class No Acknowledgement, trigger "DB302_HMI_Faults_Carrier15_Faults_3" bit 6
   1016: 'Spare_Fault_1016', class No Acknowledgement, trigger "DB302_HMI_Faults_Carrier15_Faults_3" bit 7
   1017: 'Spare_Fault_1017', class No Acknowledgement, trigger "DB302_HMI_Faults_Carrier15_Faults_3" bit 8
   1018: 'Spare_Fault_1018', class No Acknowledgement, trigger "DB302_HMI_Faults_Carrier15_Faults_3" bit 9
   1019: 'Spare_Fault_1019', class No Acknowledgement, trigger "DB302_HMI_Faults_Carrier15_Faults_3" bit 10
   1020: 'Spare_Fault_1020', class No Acknowledgement, trigger "DB302_HMI_Faults_Carrier15_Faults_3" bit 11
   1021: 'Spare_Fault_1021', class No Acknowledgement, trigger "DB302_HMI_Faults_Carrier15_Faults_3" bit 12
   1022: 'Spare_Fault_1022', class No Acknowledgement, trigger "DB302_HMI_Faults_Carrier15_Faults_3" bit 13
   1023: 'Spare_Fault_1023', class No Acknowledgement, trigger "DB302_HMI_Faults_Carrier15_Faults_3" bit 14
   1024: 'Spare_Fault_1024', class No Acknowledgement, trigger "DB302_HMI_Faults_Carrier15_Faults_3" bit 15
   1025: 'Carrier 16 Disconnect Open Power Fault DI11.0', class No Acknowledgement, trigger "DB302_HMI_Faults_Carrier16_Faults_0" bit 0
   1026: 'Carrier 16 Drive Profinet Comm Fault', class No Acknowledgement, trigger "DB302_HMI_Faults_Carrier16_Faults_0" bit 1
   1027: 'Carrier 16 Production Stop Not Reset', class No Acknowledgement, trigger "DB302_HMI_Faults_Carrier16_Faults_0" bit 2
   1028: 'Carrier 16 CB02122 Tripped', class No Acknowledgement, trigger "DB302_HMI_Faults_Carrier16_Faults_0" bit 3
   1029: 'Carrier 16 CB02123 Tripped', class No Acknowledgement, trigger "DB302_HMI_Faults_Carrier16_Faults_0" bit 4
   1030: 'Carrier 16 AUX1 CB Tripped', class No Acknowledgement, trigger "DB302_HMI_Faults_Carrier16_Faults_0" bit 5
   1031: 'Carrier 16 AUX2 CB Tripped', class No Acknowledgement, trigger "DB302_HMI_Faults_Carrier16_Faults_0" bit 6
   1032: 'Carrier 16 PLC Not Communicating', class No Acknowledgement, trigger "DB302_HMI_Faults_Carrier16_Faults_0" bit 7
   1033: 'Carrier 16 Safe Input Card Fault', class No Acknowledgement, trigger "DB302_HMI_Faults_Carrier16_Faults_0" bit 8
   1034: 'Carrier 16 Safe Output Card Fault', class No Acknowledgement, trigger "DB302_HMI_Faults_Carrier16_Faults_0" bit 9
   1035: 'Carrier 16 Standard Input Card Fault', class No Acknowledgement, trigger "DB302_HMI_Faults_Carrier16_Faults_0" bit 10
   1036: 'Carrier 16 Standard Output Card Fault', class No Acknowledgement, trigger "DB302_HMI_Faults_Carrier16_Faults_0" bit 11
   1037: 'Carrier 16 Encoder Position Fault', class No Acknowledgement, trigger "DB302_HMI_Faults_Carrier16_Faults_0" bit 12
   1038: 'Carrier 16 Encoder Internal Error', class No Acknowledgement, trigger "DB302_HMI_Faults_Carrier16_Faults_0" bit 13
   1039: 'Carrier 16 Encoder Comm Fault', class No Acknowledgement, trigger "DB302_HMI_Faults_Carrier16_Faults_0" bit 14
   1040: 'Carrier 16 HMI Comm Fault', class No Acknowledgement, trigger "DB302_HMI_Faults_Carrier16_Faults_0" bit 15
   1041: 'Carrier 16 Crash Detection Fault', class No Acknowledgement, trigger "DB302_HMI_Faults_Carrier16_Faults_1" bit 0
   1042: 'Carrier 16 Carrier Number Invalid', class No Acknowledgement, trigger "DB302_HMI_Faults_Carrier16_Faults_1" bit 1
   1043: 'Carrier 16 Drive: PROFINET configuration error', class No Acknowledgement, trigger "DB302_HMI_Faults_Carrier16_Faults_1" bit 2
   1044: 'Carrier 16 Drive: Error internal communications', class No Acknowledgement, trigger "DB302_HMI_Faults_Carrier16_Faults_1" bit 3
   1045: 'Carrier 16 Drive: Motor overtemperature', class No Acknowledgement, trigger "DB302_HMI_Faults_Carrier16_Faults_1" bit 4
   1046: 'Carrier 16 Drive: Motor overcurrent', class No Acknowledgement, trigger "DB302_HMI_Faults_Carrier16_Faults_1" bit 5
   1047: 'Carrier 16 Drive: Infeed or power unit not ready', class No Acknowledgement, trigger "DB302_HMI_Faults_Carrier16_Faults_1" bit 6
   1048: 'Carrier 16 Drive: Short-circuit/ground fault detected', class No Acknowledgement, trigger "DB302_HMI_Faults_Carrier16_Faults_1" bit 7
   1049: 'Carrier 16 Drive: PROFINET Setpoint timeout', class No Acknowledgement, trigger "DB302_HMI_Faults_Carrier16_Faults_1" bit 8
   1050: 'Carrier 16 Power unit: Overcurrent', class No Acknowledgement, trigger "DB302_HMI_Faults_Carrier16_Faults_1" bit 9
   1051: 'Carrier 16 Power unit: DC link voltage overvoltage', class No Acknowledgement, trigger "DB302_HMI_Faults_Carrier16_Faults_1" bit 10
   1052: 'Carrier 16 Power unit: DC link voltage undervoltage', class No Acknowledgement, trigger "DB302_HMI_Faults_Carrier16_Faults_1" bit 11
   1053: 'Carrier 16 Power unit: Line phase failure in main circuit', class No Acknowledgement, trigger "DB302_HMI_Faults_Carrier16_Faults_1" bit 12
   1054: 'Carrier 16 Power unit: Phase failure motor cable', class No Acknowledgement, trigger "DB302_HMI_Faults_Carrier16_Faults_1" bit 13
   1055: 'Carrier 16 Power unit: Ground fault', class No Acknowledgement, trigger "DB302_HMI_Faults_Carrier16_Faults_1" bit 14
   1056: 'Spare_Fault_1056', class No Acknowledgement, trigger "DB302_HMI_Faults_Carrier16_Faults_1" bit 15
   1057: 'Carrier 16 Motion Off Fault', class No Acknowledgement, trigger "DB302_HMI_Faults_Carrier16_Faults_2" bit 0
   1058: 'Carrier 16 Motion On Fault', class No Acknowledgement, trigger "DB302_HMI_Faults_Carrier16_Faults_2" bit 1
   1059: 'Carrier 16 Spacing Fault', class No Acknowledgement, trigger "DB302_HMI_Faults_Carrier16_Faults_2" bit 2
   1060: 'Carrier 16 Duplicate Carrier Number Fault', class No Acknowledgement, trigger "DB302_HMI_Faults_Carrier16_Faults_2" bit 3
   1061: 'Spare_Fault_1061', class No Acknowledgement, trigger "DB302_HMI_Faults_Carrier16_Faults_2" bit 4
   1062: 'Spare_Fault_1062', class No Acknowledgement, trigger "DB302_HMI_Faults_Carrier16_Faults_2" bit 5
   1063: 'Spare_Fault_1063', class No Acknowledgement, trigger "DB302_HMI_Faults_Carrier16_Faults_2" bit 6
   1064: 'Spare_Fault_1064', class No Acknowledgement, trigger "DB302_HMI_Faults_Carrier16_Faults_2" bit 7
   1065: 'Spare_Fault_1065', class No Acknowledgement, trigger "DB302_HMI_Faults_Carrier16_Faults_2" bit 8
   1066: 'Spare_Fault_1066', class No Acknowledgement, trigger "DB302_HMI_Faults_Carrier16_Faults_2" bit 9
   1067: 'Spare_Fault_1067', class No Acknowledgement, trigger "DB302_HMI_Faults_Carrier16_Faults_2" bit 10
   1068: 'Spare_Fault_1068', class No Acknowledgement, trigger "DB302_HMI_Faults_Carrier16_Faults_2" bit 11
   1069: 'Spare_Fault_1069', class No Acknowledgement, trigger "DB302_HMI_Faults_Carrier16_Faults_2" bit 12
   1070: 'Spare_Fault_1070', class No Acknowledgement, trigger "DB302_HMI_Faults_Carrier16_Faults_2" bit 13
   1071: 'Spare_Fault_1071', class No Acknowledgement, trigger "DB302_HMI_Faults_Carrier16_Faults_2" bit 14
   1072: 'Spare_Fault_1072', class No Acknowledgement, trigger "DB302_HMI_Faults_Carrier16_Faults_2" bit 15
   1073: 'Spare_Fault_1073', class No Acknowledgement, trigger "DB302_HMI_Faults_Carrier16_Faults_3" bit 0
   1074: 'Spare_Fault_1074', class No Acknowledgement, trigger "DB302_HMI_Faults_Carrier16_Faults_3" bit 1
   1075: 'Spare_Fault_1075', class No Acknowledgement, trigger "DB302_HMI_Faults_Carrier16_Faults_3" bit 2
   1076: 'Spare_Fault_1076', class No Acknowledgement, trigger "DB302_HMI_Faults_Carrier16_Faults_3" bit 3
   1077: 'Spare_Fault_1077', class No Acknowledgement, trigger "DB302_HMI_Faults_Carrier16_Faults_3" bit 4
   1078: 'Spare_Fault_1078', class No Acknowledgement, trigger "DB302_HMI_Faults_Carrier16_Faults_3" bit 5
   1079: 'Spare_Fault_1079', class No Acknowledgement, trigger "DB302_HMI_Faults_Carrier16_Faults_3" bit 6
   1080: 'Spare_Fault_1080', class No Acknowledgement, trigger "DB302_HMI_Faults_Carrier16_Faults_3" bit 7
   1081: 'Spare_Fault_1081', class No Acknowledgement, trigger "DB302_HMI_Faults_Carrier16_Faults_3" bit 8
   1082: 'Spare_Fault_1082', class No Acknowledgement, trigger "DB302_HMI_Faults_Carrier16_Faults_3" bit 9
   1083: 'Spare_Fault_1083', class No Acknowledgement, trigger "DB302_HMI_Faults_Carrier16_Faults_3" bit 10
   1084: 'Spare_Fault_1084', class No Acknowledgement, trigger "DB302_HMI_Faults_Carrier16_Faults_3" bit 11
   1085: 'Spare_Fault_1085', class No Acknowledgement, trigger "DB302_HMI_Faults_Carrier16_Faults_3" bit 12
   1086: 'Spare_Fault_1086', class No Acknowledgement, trigger "DB302_HMI_Faults_Carrier16_Faults_3" bit 13
   1087: 'Spare_Fault_1087', class No Acknowledgement, trigger "DB302_HMI_Faults_Carrier16_Faults_3" bit 14
   1088: 'Spare_Fault_1088', class No Acknowledgement, trigger "DB302_HMI_Faults_Carrier16_Faults_3" bit 15
   1089: 'Carrier 17 Disconnect Open Power Fault DI11.0', class No Acknowledgement, trigger "DB302_HMI_Faults_Carrier17_Faults_0" bit 0
   1090: 'Carrier 17 Drive Profinet Comm Fault', class No Acknowledgement, trigger "DB302_HMI_Faults_Carrier17_Faults_0" bit 1
   1091: 'Carrier 17 Production Stop Not Reset', class No Acknowledgement, trigger "DB302_HMI_Faults_Carrier17_Faults_0" bit 2
   1092: 'Carrier 17 CB02122 Tripped', class No Acknowledgement, trigger "DB302_HMI_Faults_Carrier17_Faults_0" bit 3
   1093: 'Carrier 17 CB02123 Tripped', class No Acknowledgement, trigger "DB302_HMI_Faults_Carrier17_Faults_0" bit 4
   1094: 'Carrier 17 AUX1 CB Tripped', class No Acknowledgement, trigger "DB302_HMI_Faults_Carrier17_Faults_0" bit 5
   1095: 'Carrier 17 AUX2 CB Tripped', class No Acknowledgement, trigger "DB302_HMI_Faults_Carrier17_Faults_0" bit 6
   1096: 'Carrier 17 PLC Not Communicating', class No Acknowledgement, trigger "DB302_HMI_Faults_Carrier17_Faults_0" bit 7
   1097: 'Carrier 17 Safe Input Card Fault', class No Acknowledgement, trigger "DB302_HMI_Faults_Carrier17_Faults_0" bit 8
   1098: 'Carrier 17 Safe Output Card Fault', class No Acknowledgement, trigger "DB302_HMI_Faults_Carrier17_Faults_0" bit 9
   1099: 'Carrier 17 Standard Input Card Fault', class No Acknowledgement, trigger "DB302_HMI_Faults_Carrier17_Faults_0" bit 10
   1100: 'Carrier 17 Standard Output Card Fault', class No Acknowledgement, trigger "DB302_HMI_Faults_Carrier17_Faults_0" bit 11
   1101: 'Carrier 17 Encoder Position Fault', class No Acknowledgement, trigger "DB302_HMI_Faults_Carrier17_Faults_0" bit 12
   1102: 'Carrier 17 Encoder Internal Error', class No Acknowledgement, trigger "DB302_HMI_Faults_Carrier17_Faults_0" bit 13
   1103: 'Carrier 17 Encoder Comm Fault', class No Acknowledgement, trigger "DB302_HMI_Faults_Carrier17_Faults_0" bit 14
   1104: 'Carrier 17 HMI Comm Fault', class No Acknowledgement, trigger "DB302_HMI_Faults_Carrier17_Faults_0" bit 15
   1105: 'Carrier 17 Crash Detection Fault', class No Acknowledgement, trigger "DB302_HMI_Faults_Carrier17_Faults_1" bit 0
   1106: 'Carrier 17 Carrier Number Invalid', class No Acknowledgement, trigger "DB302_HMI_Faults_Carrier17_Faults_1" bit 1
   1107: 'Carrier 17 Drive: PROFINET configuration error', class No Acknowledgement, trigger "DB302_HMI_Faults_Carrier17_Faults_1" bit 2
   1108: 'Carrier 17 Drive: Error internal communications', class No Acknowledgement, trigger "DB302_HMI_Faults_Carrier17_Faults_1" bit 3
   1109: 'Carrier 17 Drive: Motor overtemperature', class No Acknowledgement, trigger "DB302_HMI_Faults_Carrier17_Faults_1" bit 4
   1110: 'Carrier 17 Drive: Motor overcurrent', class No Acknowledgement, trigger "DB302_HMI_Faults_Carrier17_Faults_1" bit 5
   1111: 'Carrier 17 Drive: Infeed or power unit not ready', class No Acknowledgement, trigger "DB302_HMI_Faults_Carrier17_Faults_1" bit 6
   1112: 'Carrier 17 Drive: Short-circuit/ground fault detected', class No Acknowledgement, trigger "DB302_HMI_Faults_Carrier17_Faults_1" bit 7
   1113: 'Carrier 17 Drive: PROFINET Setpoint timeout', class No Acknowledgement, trigger "DB302_HMI_Faults_Carrier17_Faults_1" bit 8
   1114: 'Carrier 17 Power unit: Overcurrent', class No Acknowledgement, trigger "DB302_HMI_Faults_Carrier17_Faults_1" bit 9
   1115: 'Carrier 17 Power unit: DC link voltage overvoltage', class No Acknowledgement, trigger "DB302_HMI_Faults_Carrier17_Faults_1" bit 10
   1116: 'Carrier 17 Power unit: DC link voltage undervoltage', class No Acknowledgement, trigger "DB302_HMI_Faults_Carrier17_Faults_1" bit 11
   1117: 'Carrier 17 Power unit: Line phase failure in main circuit', class No Acknowledgement, trigger "DB302_HMI_Faults_Carrier17_Faults_1" bit 12